REGION Network 1: HL.Machine in order GREEN
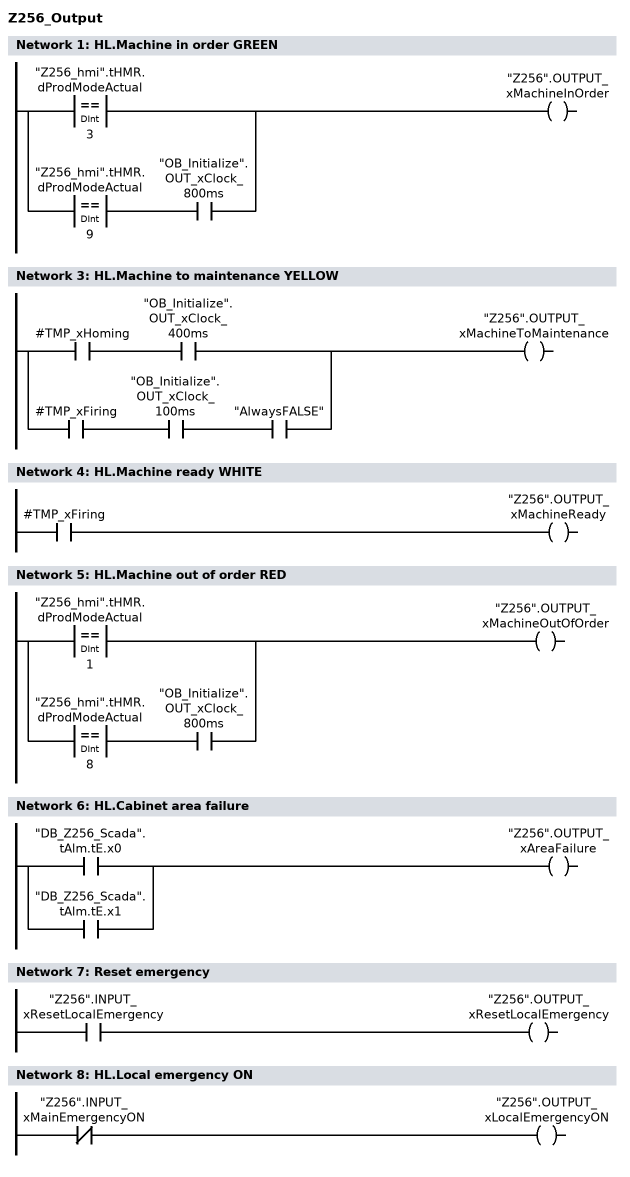
   RUNG wire#powerrail
      { S7_Templates := "SrcType := DInt" } EQ_Contact(in1 := "Z256_hmi".tHMR.dProdModeActual, in2 := 3)
      wire#w1
      Coil( "Z256".OUTPUT_xMachineInOrder )
   END_RUNG
   RUNG wire#powerrail
      { S7_Templates := "SrcType := DInt" } EQ_Contact(in1 := "Z256_hmi".tHMR.dProdModeActual, in2 := 9)
      Contact( "OB_Initialize".OUT_xClock_800ms )
   END_RUNG wire#w1
   // the same network as SCL:
   "Z256".OUTPUT_xMachineInOrder := ("Z256_hmi".tHMR.dProdModeActual = 3) OR (("Z256_hmi".tHMR.dProdModeActual = 9) AND "OB_Initialize".OUT_xClock_800ms);
END_REGION

REGION Network 2 (SCL): Homing/firing in progress
   #TMP_xHoming := false;
   #TMP_xFiring := false;
   FOR #TMP_dIndex := 0 TO "CONST_dNumberOfHeadsCycle" DO
       IF "M256_Manag_IDB".M256M_IDB[#TMP_dIndex].PH_xHeadHomeSwitch THEN
           #TMP_xHoming := true;
       END_IF;
       IF "M256_Manag_IDB".M256F_IDB[#TMP_dIndex].OUTPUT_xFireON THEN
           #TMP_xFiring := true;
       END_IF;
   END_FOR;
END_REGION

REGION Network 3: HL.Machine to maintenance YELLOW
   RUNG wire#powerrail
      Contact( #TMP_xHoming )
      Contact( "OB_Initialize".OUT_xClock_400ms )
      wire#w1
      Coil( "Z256".OUTPUT_xMachineToMaintenance )
   END_RUNG
   RUNG wire#powerrail
      Contact( #TMP_xFiring )
      Contact( "OB_Initialize".OUT_xClock_100ms )
      Contact( "AlwaysFALSE" )
   END_RUNG wire#w1
   // the same network as SCL:
   "Z256".OUTPUT_xMachineToMaintenance := (#TMP_xHoming AND "OB_Initialize".OUT_xClock_400ms) OR (#TMP_xFiring AND "OB_Initialize".OUT_xClock_100ms AND "AlwaysFALSE");
END_REGION

REGION Network 4: HL.Machine ready WHITE
   RUNG wire#powerrail
      Contact( #TMP_xFiring )
      Coil( "Z256".OUTPUT_xMachineReady )
   END_RUNG
   // the same network as SCL:
   "Z256".OUTPUT_xMachineReady := #TMP_xFiring;
END_REGION

REGION Network 5: HL.Machine out of order RED
   RUNG wire#powerrail
      { S7_Templates := "SrcType := DInt" } EQ_Contact(in1 := "Z256_hmi".tHMR.dProdModeActual, in2 := 1)
      wire#w1
      Coil( "Z256".OUTPUT_xMachineOutOfOrder )
   END_RUNG
   RUNG wire#powerrail
      { S7_Templates := "SrcType := DInt" } EQ_Contact(in1 := "Z256_hmi".tHMR.dProdModeActual, in2 := 8)
      Contact( "OB_Initialize".OUT_xClock_800ms )
   END_RUNG wire#w1
   // the same network as SCL:
   "Z256".OUTPUT_xMachineOutOfOrder := ("Z256_hmi".tHMR.dProdModeActual = 1) OR (("Z256_hmi".tHMR.dProdModeActual = 8) AND "OB_Initialize".OUT_xClock_800ms);
END_REGION

REGION Network 6: HL.Cabinet area failure
   RUNG wire#powerrail
      Contact( "DB_Z256_Scada".tAlm.tE.x0 )
      wire#w1
      Coil( "Z256".OUTPUT_xAreaFailure )
   END_RUNG
   RUNG wire#powerrail
      Contact( "DB_Z256_Scada".tAlm.tE.x1 )
   END_RUNG wire#w1
   // the same network as SCL:
   "Z256".OUTPUT_xAreaFailure := "DB_Z256_Scada".tAlm.tE.x0 OR "DB_Z256_Scada".tAlm.tE.x1;
END_REGION

REGION Network 7: Reset emergency
   RUNG wire#powerrail
      Contact( "Z256".INPUT_xResetLocalEmergency )
      Coil( "Z256".OUTPUT_xResetLocalEmergency )
   END_RUNG
   // the same network as SCL:
   "Z256".OUTPUT_xResetLocalEmergency := "Z256".INPUT_xResetLocalEmergency;
END_REGION

REGION Network 8: HL.Local emergency ON
   RUNG wire#powerrail
      I_Contact( "Z256".INPUT_xMainEmergencyON )
      Coil( "Z256".OUTPUT_xLocalEmergencyON )
   END_RUNG
   // the same network as SCL:
   "Z256".OUTPUT_xLocalEmergencyON := NOT "Z256".INPUT_xMainEmergencyON;
END_REGION

REGION Network 9 (SCL): In production selector lamp

   FOR #TMP_dIndex := 0 TO "CONST_dNumberOfHeadsCycle" DO
       IF "Z256_hmi".tHMR.rgdHeadsActualStatus[#TMP_dIndex]=3 OR ("Z256_hmi".tHMR.dProdModeActual=3 AND "OB_Initialize".OUT_xClock_800ms) THEN
           "Z256".OUTPUT_rgxHeadsInProduction[#TMP_dIndex] := true;
       ELSE
           "Z256".OUTPUT_rgxHeadsInProduction[#TMP_dIndex] := false;
       END_IF;
   END_FOR;
END_REGION
END_FUNCTION

FUNCTION "INIT_PlantCostants" : Void   // FC20, SCL
{ S7_Optimized_Access := 'TRUE' }
VERSION : 0.1
BEGIN
   //********** FOLLOW HERE THE PLANT CONSTANTS *********


   //ONLY FOR ONE LITE PLANT (when num of lites selection isn't present on scada):
   //"Z256_HMI".tHMW.dNumberOfLites := 1;


   //Connection data head #1
   "M256_Manag_IDB".IN_tConnectionData[0].ConnectID1 := 1;
   "M256_Manag_IDB".IN_tConnectionData[0].ConnectID2 := 2;
   "M256_Manag_IDB".IN_tConnectionData[0].ConnectID3 := 3;
   "M256_Manag_IDB".IN_tConnectionData[0].ConnectID4 := 4;
   "M256_Manag_IDB".IN_tConnectionData[0].IP_OCTET_1 := 192;
   "M256_Manag_IDB".IN_tConnectionData[0].IP_OCTET_2 := 168;
   "M256_Manag_IDB".IN_tConnectionData[0].IP_OCTET_3 := 22;
   "M256_Manag_IDB".IN_tConnectionData[0].IP_OCTET_4 := 21;
   //Connection data head #2
   "M256_Manag_IDB".IN_tConnectionData[1].ConnectID1 := 5;
   "M256_Manag_IDB".IN_tConnectionData[1].ConnectID2 := 6;
   "M256_Manag_IDB".IN_tConnectionData[1].ConnectID3 := 7;
   "M256_Manag_IDB".IN_tConnectionData[1].ConnectID4 := 8;
   "M256_Manag_IDB".IN_tConnectionData[1].IP_OCTET_1 := 192;
   "M256_Manag_IDB".IN_tConnectionData[1].IP_OCTET_2 := 168;
   "M256_Manag_IDB".IN_tConnectionData[1].IP_OCTET_3 := 22;
   "M256_Manag_IDB".IN_tConnectionData[1].IP_OCTET_4 := 31;
   //Connection data head #3
   "M256_Manag_IDB".IN_tConnectionData[2].ConnectID1 := 9;
   "M256_Manag_IDB".IN_tConnectionData[2].ConnectID2 := 10;
   "M256_Manag_IDB".IN_tConnectionData[2].ConnectID3 := 11;
   "M256_Manag_IDB".IN_tConnectionData[2].ConnectID4 := 12;
   "M256_Manag_IDB".IN_tConnectionData[2].IP_OCTET_1 := 192;
   "M256_Manag_IDB".IN_tConnectionData[2].IP_OCTET_2 := 168;
   "M256_Manag_IDB".IN_tConnectionData[2].IP_OCTET_3 := 22;
   "M256_Manag_IDB".IN_tConnectionData[2].IP_OCTET_4 := 51;
   //Connection data head #4
   "M256_Manag_IDB".IN_tConnectionData[3].ConnectID1 := 13;
   "M256_Manag_IDB".IN_tConnectionData[3].ConnectID2 := 14;
   "M256_Manag_IDB".IN_tConnectionData[3].ConnectID3 := 15;
   "M256_Manag_IDB".IN_tConnectionData[3].ConnectID4 := 16;
   "M256_Manag_IDB".IN_tConnectionData[3].IP_OCTET_1 := 192;
   "M256_Manag_IDB".IN_tConnectionData[3].IP_OCTET_2 := 168;
   "M256_Manag_IDB".IN_tConnectionData[3].IP_OCTET_3 := 22;
   "M256_Manag_IDB".IN_tConnectionData[3].IP_OCTET_4 := 26;

   //Connection data head #5
   "M256_Manag_IDB".IN_tConnectionData[4].ConnectID1 := 17;
   "M256_Manag_IDB".IN_tConnectionData[4].ConnectID2 := 18;
   "M256_Manag_IDB".IN_tConnectionData[4].ConnectID3 := 19;
   "M256_Manag_IDB".IN_tConnectionData[4].ConnectID4 := 20;
   "M256_Manag_IDB".IN_tConnectionData[4].IP_OCTET_1 := 192;
   "M256_Manag_IDB".IN_tConnectionData[4].IP_OCTET_2 := 168;
   "M256_Manag_IDB".IN_tConnectionData[4].IP_OCTET_3 := 22;
   "M256_Manag_IDB".IN_tConnectionData[4].IP_OCTET_4 := 35;

   //Connection data head #6
   "M256_Manag_IDB".IN_tConnectionData[4].ConnectID1 := 21;
   "M256_Manag_IDB".IN_tConnectionData[4].ConnectID2 := 22;
   "M256_Manag_IDB".IN_tConnectionData[4].ConnectID3 := 23;
   "M256_Manag_IDB".IN_tConnectionData[4].ConnectID4 := 24;
   "M256_Manag_IDB".IN_tConnectionData[4].IP_OCTET_1 := 192;
   "M256_Manag_IDB".IN_tConnectionData[4].IP_OCTET_2 := 168;
   "M256_Manag_IDB".IN_tConnectionData[4].IP_OCTET_3 := 22;
   "M256_Manag_IDB".IN_tConnectionData[4].IP_OCTET_4 := 56;

   //Connection data head #7
   "M256_Manag_IDB".IN_tConnectionData[4].ConnectID1 := 25;
   "M256_Manag_IDB".IN_tConnectionData[4].ConnectID2 := 26;
   "M256_Manag_IDB".IN_tConnectionData[4].ConnectID3 := 27;
   "M256_Manag_IDB".IN_tConnectionData[4].ConnectID4 := 28;
   "M256_Manag_IDB".IN_tConnectionData[4].IP_OCTET_1 := 192;
   "M256_Manag_IDB".IN_tConnectionData[4].IP_OCTET_2 := 168;
   "M256_Manag_IDB".IN_tConnectionData[4].IP_OCTET_3 := 22;
   "M256_Manag_IDB".IN_tConnectionData[4].IP_OCTET_4 := 46;

   //Connection data head #8
   "M256_Manag_IDB".IN_tConnectionData[4].ConnectID1 := 29;
   "M256_Manag_IDB".IN_tConnectionData[4].ConnectID2 := 30;
   "M256_Manag_IDB".IN_tConnectionData[4].ConnectID3 := 31;
   "M256_Manag_IDB".IN_tConnectionData[4].ConnectID4 := 32;
   "M256_Manag_IDB".IN_tConnectionData[4].IP_OCTET_1 := 192;
   "M256_Manag_IDB".IN_tConnectionData[4].IP_OCTET_2 := 168;
   "M256_Manag_IDB".IN_tConnectionData[4].IP_OCTET_3 := 22;
   "M256_Manag_IDB".IN_tConnectionData[4].IP_OCTET_4 := 41;

   //Operator side encumbrance operator side - Heads [mm/100]
   "PLANT_CONSTANTS".CONST_dHOpSideEnc_cmm[0] := 9500;
   "PLANT_CONSTANTS".CONST_dHOpSideEnc_cmm[1] := 2000;
   "PLANT_CONSTANTS".CONST_dHOpSideEnc_cmm[2] := 9500;
   "PLANT_CONSTANTS".CONST_dHOpSideEnc_cmm[3] := 9500;
   "PLANT_CONSTANTS".CONST_dHOpSideEnc_cmm[4] := 9500;
   "PLANT_CONSTANTS".CONST_dHOpSideEnc_cmm[5] := 9500;
   "PLANT_CONSTANTS".CONST_dHOpSideEnc_cmm[6] := 9500;
   "PLANT_CONSTANTS".CONST_dHOpSideEnc_cmm[7] := 2000;

   //Opposite operator side encumbrance - Heads [mm/100]
   "PLANT_CONSTANTS".CONST_dHOppoSideEnc_cmm[0] := 2000;
   "PLANT_CONSTANTS".CONST_dHOppoSideEnc_cmm[1] := 9500;
   "PLANT_CONSTANTS".CONST_dHOppoSideEnc_cmm[2] := 2000;
   "PLANT_CONSTANTS".CONST_dHOppoSideEnc_cmm[3] := 2000;
   "PLANT_CONSTANTS".CONST_dHOppoSideEnc_cmm[4] := 2000;
   "PLANT_CONSTANTS".CONST_dHOppoSideEnc_cmm[5] := 2000;
   "PLANT_CONSTANTS".CONST_dHOppoSideEnc_cmm[6] := 2000;
   "PLANT_CONSTANTS".CONST_dHOppoSideEnc_cmm[7] := 9500;

   //Home side
   "PLANT_CONSTANTS".CONST_rgxHomeSide[0] := 0;
   "PLANT_CONSTANTS".CONST_rgxHomeSide[1] := 0;
   "PLANT_CONSTANTS".CONST_rgxHomeSide[2] := 0;
   "PLANT_CONSTANTS".CONST_rgxHomeSide[3] := 0;
   "PLANT_CONSTANTS".CONST_rgxHomeSide[4] := 1;
   "PLANT_CONSTANTS".CONST_rgxHomeSide[5] := 1;
   "PLANT_CONSTANTS".CONST_rgxHomeSide[6] := 1;
   "PLANT_CONSTANTS".CONST_rgxHomeSide[7] := 1;

   //Pressure increment timer
   "M256_Manag_IDB".M256F_IDB[0].AUX_tmON_PressureInc.PT := t#500ms;
   "M256_Manag_IDB".M256F_IDB[1].AUX_tmON_PressureInc.PT := t#500ms;
   "M256_Manag_IDB".M256F_IDB[2].AUX_tmON_PressureInc.PT := t#500ms;
   "M256_Manag_IDB".M256F_IDB[3].AUX_tmON_PressureInc.PT := t#500ms;
   "M256_Manag_IDB".M256F_IDB[4].AUX_tmON_PressureInc.PT := t#500ms;
   "M256_Manag_IDB".M256F_IDB[5].AUX_tmON_PressureInc.PT := t#500ms;
   "M256_Manag_IDB".M256F_IDB[6].AUX_tmON_PressureInc.PT := t#500ms;
   "M256_Manag_IDB".M256F_IDB[7].AUX_tmON_PressureInc.PT := t#500ms;

   //Pressure decrement timer
   "M256_Manag_IDB".M256F_IDB[0].AUX_tmON_PressureDec.PT := t#500ms;
   "M256_Manag_IDB".M256F_IDB[1].AUX_tmON_PressureDec.PT := t#500ms;
   "M256_Manag_IDB".M256F_IDB[2].AUX_tmON_PressureDec.PT := t#500ms;
   "M256_Manag_IDB".M256F_IDB[3].AUX_tmON_PressureDec.PT := t#500ms;
   "M256_Manag_IDB".M256F_IDB[4].AUX_tmON_PressureDec.PT := t#500ms;
   "M256_Manag_IDB".M256F_IDB[5].AUX_tmON_PressureDec.PT := t#500ms;
   "M256_Manag_IDB".M256F_IDB[6].AUX_tmON_PressureDec.PT := t#500ms;
   "M256_Manag_IDB".M256F_IDB[7].AUX_tmON_PressureDec.PT := t#500ms;

   //Time head in position filters values [ms]
   "M256_Manag_IDB".M256A_IDB[0].AUX_tmON_FaultsCarrPos.PT := t#100ms;
   "M256_Manag_IDB".M256A_IDB[1].AUX_tmON_FaultsCarrPos.PT := t#100ms;
   "M256_Manag_IDB".M256A_IDB[2].AUX_tmON_FaultsCarrPos.PT := t#100ms;
   "M256_Manag_IDB".M256A_IDB[3].AUX_tmON_FaultsCarrPos.PT := t#100ms;
   "M256_Manag_IDB".M256A_IDB[4].AUX_tmON_FaultsCarrPos.PT := t#100ms;
   "M256_Manag_IDB".M256A_IDB[5].AUX_tmON_FaultsCarrPos.PT := t#100ms;
   "M256_Manag_IDB".M256A_IDB[6].AUX_tmON_FaultsCarrPos.PT := t#100ms;
   "M256_Manag_IDB".M256A_IDB[7].AUX_tmON_FaultsCarrPos.PT := t#100ms;

   "M256_Manag_IDB".M256A_IDB[0].AUX_tmOFF_FaultsCarrPos.PT := t#100ms;
   "M256_Manag_IDB".M256A_IDB[1].AUX_tmOFF_FaultsCarrPos.PT := t#100ms;
   "M256_Manag_IDB".M256A_IDB[2].AUX_tmOFF_FaultsCarrPos.PT := t#100ms;
   "M256_Manag_IDB".M256A_IDB[3].AUX_tmOFF_FaultsCarrPos.PT := t#100ms;
   "M256_Manag_IDB".M256A_IDB[4].AUX_tmOFF_FaultsCarrPos.PT := t#100ms;
   "M256_Manag_IDB".M256A_IDB[5].AUX_tmOFF_FaultsCarrPos.PT := t#100ms;
   "M256_Manag_IDB".M256A_IDB[6].AUX_tmOFF_FaultsCarrPos.PT := t#100ms;
   "M256_Manag_IDB".M256A_IDB[7].AUX_tmOFF_FaultsCarrPos.PT := t#100ms;

   //Timer driver enable retain
   "M256_Manag_IDB".M256M_IDB[0].AUX_tmDriveReadyRetainTimer.PT := t#100ms;
   "M256_Manag_IDB".M256M_IDB[1].AUX_tmDriveReadyRetainTimer.PT := t#100ms;
   "M256_Manag_IDB".M256M_IDB[2].AUX_tmDriveReadyRetainTimer.PT := t#100ms;
   "M256_Manag_IDB".M256M_IDB[3].AUX_tmDriveReadyRetainTimer.PT := t#100ms;
   "M256_Manag_IDB".M256M_IDB[4].AUX_tmDriveReadyRetainTimer.PT := t#100ms;
   "M256_Manag_IDB".M256M_IDB[5].AUX_tmDriveReadyRetainTimer.PT := t#100ms;
   "M256_Manag_IDB".M256M_IDB[6].AUX_tmDriveReadyRetainTimer.PT := t#100ms;
   "M256_Manag_IDB".M256M_IDB[7].AUX_tmDriveReadyRetainTimer.PT := t#100ms;


   //Timer driver in movement
   "M256_Manag_IDB".M256M_IDB[0].AUX_tmOFFDriveEnable.PT := t#500ms;
   "M256_Manag_IDB".M256M_IDB[1].AUX_tmOFFDriveEnable.PT := t#500ms;
   "M256_Manag_IDB".M256M_IDB[2].AUX_tmOFFDriveEnable.PT := t#500ms;
   "M256_Manag_IDB".M256M_IDB[3].AUX_tmOFFDriveEnable.PT := t#500ms;
   "M256_Manag_IDB".M256M_IDB[4].AUX_tmOFFDriveEnable.PT := t#500ms;
   "M256_Manag_IDB".M256M_IDB[5].AUX_tmOFFDriveEnable.PT := t#500ms;
   "M256_Manag_IDB".M256M_IDB[6].AUX_tmOFFDriveEnable.PT := t#500ms;
   "M256_Manag_IDB".M256M_IDB[7].AUX_tmOFFDriveEnable.PT := t#500ms;

   "M256_Manag_IDB".M256M_IDB[0].AUX_tmOFFEnablePositioningAfterHome.PT := t#4s;
   "M256_Manag_IDB".M256M_IDB[1].AUX_tmOFFEnablePositioningAfterHome.PT := t#4s;
   "M256_Manag_IDB".M256M_IDB[2].AUX_tmOFFEnablePositioningAfterHome.PT := t#4s;
   "M256_Manag_IDB".M256M_IDB[3].AUX_tmOFFEnablePositioningAfterHome.PT := t#4s;
   "M256_Manag_IDB".M256M_IDB[4].AUX_tmOFFEnablePositioningAfterHome.PT := t#4s;
   "M256_Manag_IDB".M256M_IDB[5].AUX_tmOFFEnablePositioningAfterHome.PT := t#4s;
   "M256_Manag_IDB".M256M_IDB[6].AUX_tmOFFEnablePositioningAfterHome.PT := t#4s;
   "M256_Manag_IDB".M256M_IDB[7].AUX_tmOFFEnablePositioningAfterHome.PT := t#4s;
   //-------------HEAD #1 PARAMETERS--------------------------

   "PLANT_CONSTANTS".CONST_rgtHeadPar[0].dParametersToDownload := 17;

   //Parameter IOfunct_LIO1
   "PLANT_CONSTANTS".CONST_rgtHeadPar[0].rgtAxisParameters[0].iAddress := 1826;
   "PLANT_CONSTANTS".CONST_rgtHeadPar[0].rgtAxisParameters[0].iLength := 2;
   "PLANT_CONSTANTS".CONST_rgtHeadPar[0].rgtAxisParameters[0].dValue := 20;

   //Parameter IOfunct_LIO2
   "PLANT_CONSTANTS".CONST_rgtHeadPar[0].rgtAxisParameters[1].iAddress := 1828;
   "PLANT_CONSTANTS".CONST_rgtHeadPar[0].rgtAxisParameters[1].iLength := 2;
   "PLANT_CONSTANTS".CONST_rgtHeadPar[0].rgtAxisParameters[1].dValue := 1;

   //Parameter IOfunct_LIO3
   "PLANT_CONSTANTS".CONST_rgtHeadPar[0].rgtAxisParameters[2].iAddress := 1830;
   "PLANT_CONSTANTS".CONST_rgtHeadPar[0].rgtAxisParameters[2].iLength := 2;
   "PLANT_CONSTANTS".CONST_rgtHeadPar[0].rgtAxisParameters[2].dValue := 1;

   //Parameter IOfunct_LIO4
   "PLANT_CONSTANTS".CONST_rgtHeadPar[0].rgtAxisParameters[3].iAddress := 1832;
   "PLANT_CONSTANTS".CONST_rgtHeadPar[0].rgtAxisParameters[3].iLength := 2;
   "PLANT_CONSTANTS".CONST_rgtHeadPar[0].rgtAxisParameters[3].dValue := 1;

   //Parameter IOsigLimN
   "PLANT_CONSTANTS".CONST_rgtHeadPar[0].rgtAxisParameters[4].iAddress := 1566;
   "PLANT_CONSTANTS".CONST_rgtHeadPar[0].rgtAxisParameters[4].iLength := 2;
   "PLANT_CONSTANTS".CONST_rgtHeadPar[0].rgtAxisParameters[4].dValue := 0;

   //Parameter IOsigLimP
   "PLANT_CONSTANTS".CONST_rgtHeadPar[0].rgtAxisParameters[5].iAddress := 1568;
   "PLANT_CONSTANTS".CONST_rgtHeadPar[0].rgtAxisParameters[5].iLength := 2;
   "PLANT_CONSTANTS".CONST_rgtHeadPar[0].rgtAxisParameters[5].dValue := 0;

   //Parameter IOsigRef
   "PLANT_CONSTANTS".CONST_rgtHeadPar[0].rgtAxisParameters[6].iAddress := 1564;
   "PLANT_CONSTANTS".CONST_rgtHeadPar[0].rgtAxisParameters[6].iLength := 2;
   "PLANT_CONSTANTS".CONST_rgtHeadPar[0].rgtAxisParameters[6].dValue := 2;

   //Parameter POSdirOfRotat
   "PLANT_CONSTANTS".CONST_rgtHeadPar[0].rgtAxisParameters[7].iAddress := 1560;
   "PLANT_CONSTANTS".CONST_rgtHeadPar[0].rgtAxisParameters[7].iLength := 2;
   "PLANT_CONSTANTS".CONST_rgtHeadPar[0].rgtAxisParameters[7].dValue := 0;

   //Parameter POSscaleDenom
   "PLANT_CONSTANTS".CONST_rgtHeadPar[0].rgtAxisParameters[8].iAddress := 1550;
   "PLANT_CONSTANTS".CONST_rgtHeadPar[0].rgtAxisParameters[8].iLength := 4;
   "PLANT_CONSTANTS".CONST_rgtHeadPar[0].rgtAxisParameters[8].dValue := 500;

   //Parameter POSscaleNum
   "PLANT_CONSTANTS".CONST_rgtHeadPar[0].rgtAxisParameters[9].iAddress := 1552;
   "PLANT_CONSTANTS".CONST_rgtHeadPar[0].rgtAxisParameters[9].iLength := 4;
   "PLANT_CONSTANTS".CONST_rgtHeadPar[0].rgtAxisParameters[9].dValue := 1;

   //Parameter RAMPacc
   "PLANT_CONSTANTS".CONST_rgtHeadPar[0].rgtAxisParameters[10].iAddress := 1556;
   "PLANT_CONSTANTS".CONST_rgtHeadPar[0].rgtAxisParameters[10].iLength := 4;
   "PLANT_CONSTANTS".CONST_rgtHeadPar[0].rgtAxisParameters[10].dValue := 20000;//[rot/min]

   //Parameter RAMPdecel
   "PLANT_CONSTANTS".CONST_rgtHeadPar[0].rgtAxisParameters[11].iAddress := 1558;
   "PLANT_CONSTANTS".CONST_rgtHeadPar[0].rgtAxisParameters[11].iLength := 4;
   "PLANT_CONSTANTS".CONST_rgtHeadPar[0].rgtAxisParameters[11].dValue := 20000;//[rot/min]

   //Parameter JOGn_fast
   "PLANT_CONSTANTS".CONST_rgtHeadPar[0].rgtAxisParameters[12].iAddress := 10506;
   "PLANT_CONSTANTS".CONST_rgtHeadPar[0].rgtAxisParameters[12].iLength := 2;
   "PLANT_CONSTANTS".CONST_rgtHeadPar[0].rgtAxisParameters[12].dValue := 1000;//[rot/s2]

   //Parameter JOGn_slow
   "PLANT_CONSTANTS".CONST_rgtHeadPar[0].rgtAxisParameters[13].iAddress := 10504;
   "PLANT_CONSTANTS".CONST_rgtHeadPar[0].rgtAxisParameters[13].iLength := 2;
   "PLANT_CONSTANTS".CONST_rgtHeadPar[0].rgtAxisParameters[13].dValue := 1000;//[rot/s2]

   //Parameter JOGstepusr
   "PLANT_CONSTANTS".CONST_rgtHeadPar[0].rgtAxisParameters[14].iAddress := 10510;
   "PLANT_CONSTANTS".CONST_rgtHeadPar[0].rgtAxisParameters[14].iLength := 4;
   "PLANT_CONSTANTS".CONST_rgtHeadPar[0].rgtAxisParameters[14].dValue := 0;

   //Parameter JOGtime
   "PLANT_CONSTANTS".CONST_rgtHeadPar[0].rgtAxisParameters[15].iAddress := 10512;
   "PLANT_CONSTANTS".CONST_rgtHeadPar[0].rgtAxisParameters[15].iLength := 2;
   "PLANT_CONSTANTS".CONST_rgtHeadPar[0].rgtAxisParameters[15].dValue := 1;

   //Parameter PAReeprSave ---MUST BE THE LAST!!!
   "PLANT_CONSTANTS".CONST_rgtHeadPar[0].rgtAxisParameters[16].iAddress := 1026;
   "PLANT_CONSTANTS".CONST_rgtHeadPar[0].rgtAxisParameters[16].iLength := 2;
   "PLANT_CONSTANTS".CONST_rgtHeadPar[0].rgtAxisParameters[16].dValue := 1;

   //-------------HEAD #2 PARAMETERS--------------------------

   "PLANT_CONSTANTS".CONST_rgtHeadPar[1].dParametersToDownload := 17;

   //Parameter IOfunct_LIO1
   "PLANT_CONSTANTS".CONST_rgtHeadPar[1].rgtAxisParameters[0].iAddress := 1826;
   "PLANT_CONSTANTS".CONST_rgtHeadPar[1].rgtAxisParameters[0].iLength := 2;
   "PLANT_CONSTANTS".CONST_rgtHeadPar[1].rgtAxisParameters[0].dValue := 20;

   //Parameter IOfunct_LIO2
   "PLANT_CONSTANTS".CONST_rgtHeadPar[1].rgtAxisParameters[1].iAddress := 1828;
   "PLANT_CONSTANTS".CONST_rgtHeadPar[1].rgtAxisParameters[1].iLength := 2;
   "PLANT_CONSTANTS".CONST_rgtHeadPar[1].rgtAxisParameters[1].dValue := 1;

   //Parameter IOfunct_LIO3
   "PLANT_CONSTANTS".CONST_rgtHeadPar[1].rgtAxisParameters[2].iAddress := 1830;
   "PLANT_CONSTANTS".CONST_rgtHeadPar[1].rgtAxisParameters[2].iLength := 2;
   "PLANT_CONSTANTS".CONST_rgtHeadPar[1].rgtAxisParameters[2].dValue := 1;

   //Parameter IOfunct_LIO4
   "PLANT_CONSTANTS".CONST_rgtHeadPar[1].rgtAxisParameters[3].iAddress := 1832;
   "PLANT_CONSTANTS".CONST_rgtHeadPar[1].rgtAxisParameters[3].iLength := 2;
   "PLANT_CONSTANTS".CONST_rgtHeadPar[1].rgtAxisParameters[3].dValue := 1;

   //Parameter IOsigLimN
   "PLANT_CONSTANTS".CONST_rgtHeadPar[1].rgtAxisParameters[4].iAddress := 1566;
   "PLANT_CONSTANTS".CONST_rgtHeadPar[1].rgtAxisParameters[4].iLength := 2;
   "PLANT_CONSTANTS".CONST_rgtHeadPar[1].rgtAxisParameters[4].dValue := 0;

   //Parameter IOsigLimP
   "PLANT_CONSTANTS".CONST_rgtHeadPar[1].rgtAxisParameters[5].iAddress := 1568;
   "PLANT_CONSTANTS".CONST_rgtHeadPar[1].rgtAxisParameters[5].iLength := 2;
   "PLANT_CONSTANTS".CONST_rgtHeadPar[1].rgtAxisParameters[5].dValue := 0;

   //Parameter IOsigRef
   "PLANT_CONSTANTS".CONST_rgtHeadPar[1].rgtAxisParameters[6].iAddress := 1564;
   "PLANT_CONSTANTS".CONST_rgtHeadPar[1].rgtAxisParameters[6].iLength := 2;
   "PLANT_CONSTANTS".CONST_rgtHeadPar[1].rgtAxisParameters[6].dValue := 2;

   //Parameter POSdirOfRotat
   "PLANT_CONSTANTS".CONST_rgtHeadPar[1].rgtAxisParameters[7].iAddress := 1560;
   "PLANT_CONSTANTS".CONST_rgtHeadPar[1].rgtAxisParameters[7].iLength := 2;
   "PLANT_CONSTANTS".CONST_rgtHeadPar[1].rgtAxisParameters[7].dValue := 0;

   //Parameter POSscaleDenom
   "PLANT_CONSTANTS".CONST_rgtHeadPar[1].rgtAxisParameters[8].iAddress := 1550;
   "PLANT_CONSTANTS".CONST_rgtHeadPar[1].rgtAxisParameters[8].iLength := 4;
   "PLANT_CONSTANTS".CONST_rgtHeadPar[1].rgtAxisParameters[8].dValue := 500;

   //Parameter POSscaleNum
   "PLANT_CONSTANTS".CONST_rgtHeadPar[1].rgtAxisParameters[9].iAddress := 1552;
   "PLANT_CONSTANTS".CONST_rgtHeadPar[1].rgtAxisParameters[9].iLength := 4;
   "PLANT_CONSTANTS".CONST_rgtHeadPar[1].rgtAxisParameters[9].dValue := 1;

   //Parameter RAMPacc
   "PLANT_CONSTANTS".CONST_rgtHeadPar[1].rgtAxisParameters[10].iAddress := 1556;
   "PLANT_CONSTANTS".CONST_rgtHeadPar[1].rgtAxisParameters[10].iLength := 4;
   "PLANT_CONSTANTS".CONST_rgtHeadPar[1].rgtAxisParameters[10].dValue := 20000;//[rot/min]

   //Parameter RAMPdecel
   "PLANT_CONSTANTS".CONST_rgtHeadPar[1].rgtAxisParameters[11].iAddress := 1558;
   "PLANT_CONSTANTS".CONST_rgtHeadPar[1].rgtAxisParameters[11].iLength := 4;
   "PLANT_CONSTANTS".CONST_rgtHeadPar[1].rgtAxisParameters[11].dValue := 20000;//[rot/min]

   //Parameter JOGn_fast
   "PLANT_CONSTANTS".CONST_rgtHeadPar[1].rgtAxisParameters[12].iAddress := 10506;
   "PLANT_CONSTANTS".CONST_rgtHeadPar[1].rgtAxisParameters[12].iLength := 2;
   "PLANT_CONSTANTS".CONST_rgtHeadPar[1].rgtAxisParameters[12].dValue := 1000;//[rot/s2]

   //Parameter JOGn_slow
   "PLANT_CONSTANTS".CONST_rgtHeadPar[1].rgtAxisParameters[13].iAddress := 10504;
   "PLANT_CONSTANTS".CONST_rgtHeadPar[1].rgtAxisParameters[13].iLength := 2;
   "PLANT_CONSTANTS".CONST_rgtHeadPar[1].rgtAxisParameters[13].dValue := 1000;//[rot/s2]

   //Parameter JOGstepusr
   "PLANT_CONSTANTS".CONST_rgtHeadPar[1].rgtAxisParameters[14].iAddress := 10510;
   "PLANT_CONSTANTS".CONST_rgtHeadPar[1].rgtAxisParameters[14].iLength := 4;
   "PLANT_CONSTANTS".CONST_rgtHeadPar[1].rgtAxisParameters[14].dValue := 0;

   //Parameter JOGtime
   "PLANT_CONSTANTS".CONST_rgtHeadPar[1].rgtAxisParameters[15].iAddress := 10512;
   "PLANT_CONSTANTS".CONST_rgtHeadPar[1].rgtAxisParameters[15].iLength := 2;
   "PLANT_CONSTANTS".CONST_rgtHeadPar[1].rgtAxisParameters[15].dValue := 1;

   //Parameter PAReeprSave ---MUST BE THE LAST!!!
   "PLANT_CONSTANTS".CONST_rgtHeadPar[1].rgtAxisParameters[16].iAddress := 1026;
   "PLANT_CONSTANTS".CONST_rgtHeadPar[1].rgtAxisParameters[16].iLength := 2;
   "PLANT_CONSTANTS".CONST_rgtHeadPar[1].rgtAxisParameters[16].dValue := 1;

   //-------------HEAD #3 PARAMETERS--------------------------

   "PLANT_CONSTANTS".CONST_rgtHeadPar[2].dParametersToDownload := 17;

   //Parameter IOfunct_LIO1
   "PLANT_CONSTANTS".CONST_rgtHeadPar[2].rgtAxisParameters[0].iAddress := 1826;
   "PLANT_CONSTANTS".CONST_rgtHeadPar[2].rgtAxisParameters[0].iLength := 2;
   "PLANT_CONSTANTS".CONST_rgtHeadPar[2].rgtAxisParameters[0].dValue := 20;

   //Parameter IOfunct_LIO2
   "PLANT_CONSTANTS".CONST_rgtHeadPar[2].rgtAxisParameters[1].iAddress := 1828;
   "PLANT_CONSTANTS".CONST_rgtHeadPar[2].rgtAxisParameters[1].iLength := 2;
   "PLANT_CONSTANTS".CONST_rgtHeadPar[2].rgtAxisParameters[1].dValue := 1;

   //Parameter IOfunct_LIO3
   "PLANT_CONSTANTS".CONST_rgtHeadPar[2].rgtAxisParameters[2].iAddress := 1830;
   "PLANT_CONSTANTS".CONST_rgtHeadPar[2].rgtAxisParameters[2].iLength := 2;
   "PLANT_CONSTANTS".CONST_rgtHeadPar[2].rgtAxisParameters[2].dValue := 1;

   //Parameter IOfunct_LIO4
   "PLANT_CONSTANTS".CONST_rgtHeadPar[2].rgtAxisParameters[3].iAddress := 1832;
   "PLANT_CONSTANTS".CONST_rgtHeadPar[2].rgtAxisParameters[3].iLength := 2;
   "PLANT_CONSTANTS".CONST_rgtHeadPar[2].rgtAxisParameters[3].dValue := 1;

   //Parameter IOsigLimN
   "PLANT_CONSTANTS".CONST_rgtHeadPar[2].rgtAxisParameters[4].iAddress := 1566;
   "PLANT_CONSTANTS".CONST_rgtHeadPar[2].rgtAxisParameters[4].iLength := 2;
   "PLANT_CONSTANTS".CONST_rgtHeadPar[2].rgtAxisParameters[4].dValue := 0;

   //Parameter IOsigLimP
   "PLANT_CONSTANTS".CONST_rgtHeadPar[2].rgtAxisParameters[5].iAddress := 1568;
   "PLANT_CONSTANTS".CONST_rgtHeadPar[2].rgtAxisParameters[5].iLength := 2;
   "PLANT_CONSTANTS".CONST_rgtHeadPar[2].rgtAxisParameters[5].dValue := 0;

   //Parameter IOsigRef
   "PLANT_CONSTANTS".CONST_rgtHeadPar[2].rgtAxisParameters[6].iAddress := 1564;
   "PLANT_CONSTANTS".CONST_rgtHeadPar[2].rgtAxisParameters[6].iLength := 2;
   "PLANT_CONSTANTS".CONST_rgtHeadPar[2].rgtAxisParameters[6].dValue := 2;

   //Parameter POSdirOfRotat
   "PLANT_CONSTANTS".CONST_rgtHeadPar[2].rgtAxisParameters[7].iAddress := 1560;
   "PLANT_CONSTANTS".CONST_rgtHeadPar[2].rgtAxisParameters[7].iLength := 2;
   "PLANT_CONSTANTS".CONST_rgtHeadPar[2].rgtAxisParameters[7].dValue := 0;

   //Parameter POSscaleDenom
   "PLANT_CONSTANTS".CONST_rgtHeadPar[2].rgtAxisParameters[8].iAddress := 1550;
   "PLANT_CONSTANTS".CONST_rgtHeadPar[2].rgtAxisParameters[8].iLength := 4;
   "PLANT_CONSTANTS".CONST_rgtHeadPar[2].rgtAxisParameters[8].dValue := 500;

   //Parameter POSscaleNum
   "PLANT_CONSTANTS".CONST_rgtHeadPar[2].rgtAxisParameters[9].iAddress := 1552;
   "PLANT_CONSTANTS".CONST_rgtHeadPar[2].rgtAxisParameters[9].iLength := 4;
   "PLANT_CONSTANTS".CONST_rgtHeadPar[2].rgtAxisParameters[9].dValue := 1;

   //Parameter RAMPacc
   "PLANT_CONSTANTS".CONST_rgtHeadPar[2].rgtAxisParameters[10].iAddress := 1556;
   "PLANT_CONSTANTS".CONST_rgtHeadPar[2].rgtAxisParameters[10].iLength := 4;
   "PLANT_CONSTANTS".CONST_rgtHeadPar[2].rgtAxisParameters[10].dValue := 20000;//[rot/min]

   //Parameter RAMPdecel
   "PLANT_CONSTANTS".CONST_rgtHeadPar[2].rgtAxisParameters[11].iAddress := 1558;
   "PLANT_CONSTANTS".CONST_rgtHeadPar[2].rgtAxisParameters[11].iLength := 4;
   "PLANT_CONSTANTS".CONST_rgtHeadPar[2].rgtAxisParameters[11].dValue := 20000;//[rot/min]

   //Parameter JOGn_fast
   "PLANT_CONSTANTS".CONST_rgtHeadPar[2].rgtAxisParameters[12].iAddress := 10506;
   "PLANT_CONSTANTS".CONST_rgtHeadPar[2].rgtAxisParameters[12].iLength := 2;
   "PLANT_CONSTANTS".CONST_rgtHeadPar[2].rgtAxisParameters[12].dValue := 1000;//[rot/s2]

   //Parameter JOGn_slow
   "PLANT_CONSTANTS".CONST_rgtHeadPar[2].rgtAxisParameters[13].iAddress := 10504;
   "PLANT_CONSTANTS".CONST_rgtHeadPar[2].rgtAxisParameters[13].iLength := 2;
   "PLANT_CONSTANTS".CONST_rgtHeadPar[2].rgtAxisParameters[13].dValue := 1000;//[rot/s2]

   //Parameter JOGstepusr
   "PLANT_CONSTANTS".CONST_rgtHeadPar[2].rgtAxisParameters[14].iAddress := 10510;
   "PLANT_CONSTANTS".CONST_rgtHeadPar[2].rgtAxisParameters[14].iLength := 4;
   "PLANT_CONSTANTS".CONST_rgtHeadPar[2].rgtAxisParameters[14].dValue := 0;

   //Parameter JOGtime
   "PLANT_CONSTANTS".CONST_rgtHeadPar[2].rgtAxisParameters[15].iAddress := 10512;
   "PLANT_CONSTANTS".CONST_rgtHeadPar[2].rgtAxisParameters[15].iLength := 2;
   "PLANT_CONSTANTS".CONST_rgtHeadPar[2].rgtAxisParameters[15].dValue := 1;

   //Parameter PAReeprSave ---MUST BE THE LAST!!!
   "PLANT_CONSTANTS".CONST_rgtHeadPar[2].rgtAxisParameters[16].iAddress := 1026;
   "PLANT_CONSTANTS".CONST_rgtHeadPar[2].rgtAxisParameters[16].iLength := 2;
   "PLANT_CONSTANTS".CONST_rgtHeadPar[2].rgtAxisParameters[16].dValue := 1;

   //-------------HEAD #4 PARAMETERS--------------------------

   "PLANT_CONSTANTS".CONST_rgtHeadPar[3].dParametersToDownload := 17;

   //Parameter IOfunct_LIO1
   "PLANT_CONSTANTS".CONST_rgtHeadPar[3].rgtAxisParameters[0].iAddress := 1826;
   "PLANT_CONSTANTS".CONST_rgtHeadPar[3].rgtAxisParameters[0].iLength := 2;
   "PLANT_CONSTANTS".CONST_rgtHeadPar[3].rgtAxisParameters[0].dValue := 20;

   //Parameter IOfunct_LIO2
   "PLANT_CONSTANTS".CONST_rgtHeadPar[3].rgtAxisParameters[1].iAddress := 1828;
   "PLANT_CONSTANTS".CONST_rgtHeadPar[3].rgtAxisParameters[1].iLength := 2;
   "PLANT_CONSTANTS".CONST_rgtHeadPar[3].rgtAxisParameters[1].dValue := 1;

   //Parameter IOfunct_LIO3
   "PLANT_CONSTANTS".CONST_rgtHeadPar[3].rgtAxisParameters[2].iAddress := 1830;
   "PLANT_CONSTANTS".CONST_rgtHeadPar[3].rgtAxisParameters[2].iLength := 2;
   "PLANT_CONSTANTS".CONST_rgtHeadPar[3].rgtAxisParameters[2].dValue := 1;

   //Parameter IOfunct_LIO4
   "PLANT_CONSTANTS".CONST_rgtHeadPar[3].rgtAxisParameters[3].iAddress := 1832;
   "PLANT_CONSTANTS".CONST_rgtHeadPar[3].rgtAxisParameters[3].iLength := 2;
   "PLANT_CONSTANTS".CONST_rgtHeadPar[3].rgtAxisParameters[3].dValue := 1;

   //Parameter IOsigLimN
   "PLANT_CONSTANTS".CONST_rgtHeadPar[3].rgtAxisParameters[4].iAddress := 1566;
   "PLANT_CONSTANTS".CONST_rgtHeadPar[3].rgtAxisParameters[4].iLength := 2;
   "PLANT_CONSTANTS".CONST_rgtHeadPar[3].rgtAxisParameters[4].dValue := 0;

   //Parameter IOsigLimP
   "PLANT_CONSTANTS".CONST_rgtHeadPar[3].rgtAxisParameters[5].iAddress := 1568;
   "PLANT_CONSTANTS".CONST_rgtHeadPar[3].rgtAxisParameters[5].iLength := 2;
   "PLANT_CONSTANTS".CONST_rgtHeadPar[3].rgtAxisParameters[5].dValue := 0;

   //Parameter IOsigRef
   "PLANT_CONSTANTS".CONST_rgtHeadPar[3].rgtAxisParameters[6].iAddress := 1564;
   "PLANT_CONSTANTS".CONST_rgtHeadPar[3].rgtAxisParameters[6].iLength := 2;
   "PLANT_CONSTANTS".CONST_rgtHeadPar[3].rgtAxisParameters[6].dValue := 2;

   //Parameter POSdirOfRotat
   "PLANT_CONSTANTS".CONST_rgtHeadPar[3].rgtAxisParameters[7].iAddress := 1560;
   "PLANT_CONSTANTS".CONST_rgtHeadPar[3].rgtAxisParameters[7].iLength := 2;
   "PLANT_CONSTANTS".CONST_rgtHeadPar[3].rgtAxisParameters[7].dValue := 0;

   //Parameter POSscaleDenom
   "PLANT_CONSTANTS".CONST_rgtHeadPar[3].rgtAxisParameters[8].iAddress := 1550;
   "PLANT_CONSTANTS".CONST_rgtHeadPar[3].rgtAxisParameters[8].iLength := 4;
   "PLANT_CONSTANTS".CONST_rgtHeadPar[3].rgtAxisParameters[8].dValue := 500;

   //Parameter POSscaleNum
   "PLANT_CONSTANTS".CONST_rgtHeadPar[3].rgtAxisParameters[9].iAddress := 1552;
   "PLANT_CONSTANTS".CONST_rgtHeadPar[3].rgtAxisParameters[9].iLength := 4;
   "PLANT_CONSTANTS".CONST_rgtHeadPar[3].rgtAxisParameters[9].dValue := 1;

   //Parameter RAMPacc
   "PLANT_CONSTANTS".CONST_rgtHeadPar[3].rgtAxisParameters[10].iAddress := 1556;
   "PLANT_CONSTANTS".CONST_rgtHeadPar[3].rgtAxisParameters[10].iLength := 4;
   "PLANT_CONSTANTS".CONST_rgtHeadPar[3].rgtAxisParameters[10].dValue := 20000;//[rot/s2]

   //Parameter RAMPdecel
   "PLANT_CONSTANTS".CONST_rgtHeadPar[3].rgtAxisParameters[11].iAddress := 1558;
   "PLANT_CONSTANTS".CONST_rgtHeadPar[3].rgtAxisParameters[11].iLength := 4;
   "PLANT_CONSTANTS".CONST_rgtHeadPar[3].rgtAxisParameters[11].dValue := 20000;//[rot/s2]

   //Parameter JOGn_fast
   "PLANT_CONSTANTS".CONST_rgtHeadPar[3].rgtAxisParameters[12].iAddress := 10506;
   "PLANT_CONSTANTS".CONST_rgtHeadPar[3].rgtAxisParameters[12].iLength := 2;
   "PLANT_CONSTANTS".CONST_rgtHeadPar[3].rgtAxisParameters[12].dValue := 1000;//[rot/min]

   //Parameter JOGn_slow
   "PLANT_CONSTANTS".CONST_rgtHeadPar[3].rgtAxisParameters[13].iAddress := 10504;
   "PLANT_CONSTANTS".CONST_rgtHeadPar[3].rgtAxisParameters[13].iLength := 2;
   "PLANT_CONSTANTS".CONST_rgtHeadPar[3].rgtAxisParameters[13].dValue := 1000;//[rot/min]

   //Parameter JOGstepusr
   "PLANT_CONSTANTS".CONST_rgtHeadPar[3].rgtAxisParameters[14].iAddress := 10510;
   "PLANT_CONSTANTS".CONST_rgtHeadPar[3].rgtAxisParameters[14].iLength := 4;
   "PLANT_CONSTANTS".CONST_rgtHeadPar[3].rgtAxisParameters[14].dValue := 0;

   //Parameter JOGtime
   "PLANT_CONSTANTS".CONST_rgtHeadPar[3].rgtAxisParameters[15].iAddress := 10512;
   "PLANT_CONSTANTS".CONST_rgtHeadPar[3].rgtAxisParameters[15].iLength := 2;
   "PLANT_CONSTANTS".CONST_rgtHeadPar[3].rgtAxisParameters[15].dValue := 1;

   //Parameter PAReeprSave ---MUST BE THE LAST!!!
   "PLANT_CONSTANTS".CONST_rgtHeadPar[3].rgtAxisParameters[16].iAddress := 1026;
   "PLANT_CONSTANTS".CONST_rgtHeadPar[3].rgtAxisParameters[16].iLength := 2;
   "PLANT_CONSTANTS".CONST_rgtHeadPar[3].rgtAxisParameters[16].dValue := 1;